(* Logix 5000 project; controller _GigaDiscovery vendor 1 type 14 code 244 rev 35.11; software revision 35.03; part 15 of 23 *)
(* tags used below, declared in another part *)
   Brake_Delay : TIMER;
   Os : DINT;
   Timer_Loc : TIMER[50];
   All_Rack_Closed_Mem : BOOL;
   All_RESTRAINTS_Opened : BOOL;
   DC_Field_Motor_7 : UDT_CROUT;   // DC Field Motor 7 Gondola Contactor -Q16101E -Q16103E
   DC_Field_Pylon_Motors : UDT_CROUT;   // DC Field Pylon Motors Contactor -Q10101E -Q10103E
   Enable_to_Start : UDT_CROUT;   // Abilitazione allo start QC8011E QC8013E
   Girella_Field_Actuate_During_Inactivity : BOOL;
   Gondola_Drive_Enable : UDT_CROUT;   // Gondola Drive Ch1-Ch2 Start Enable Contactors -Q16105E -Q16107E
   I_EStop_Pb_OCC1 : UDT_DCI_STOP_TEST;   // +OCC E-stop -S30301F
   I_EStop_Pb_OCC2 : UDT_DCI_STOP_TEST;   // +OCC2 E-Stop -S28502F
   I_Gondola_Home_Position : BOOL;   // Gondola Home Position -B40002I -B40007I
   I_OCC2_Disable : UDT_DCM;   // OCC 2 CONTROL DISABLE Page 310
   I_OCC_LockOut_Motion : UDT_DCM;   // OCC -Lockout Motion -Q31203E
   I_OCC_Operator_Enable_Key : BOOL;   // OCC Console Enabled -S30305F
   I_Platform_Line_Unlock_Pressure_Switch : BOOL;   // Unlock Platform Line Pressure Switch -S22006B
   I_Platform_Opened : UDT_DCM;   // Platform Opened RFID Series -Q23801J -Q23807J
   I_Platform_Pressure_on_Close_Circuit : BOOL;   // Platform Maximum Closing Pressure -S21510B
   No_Sfty : Std_to_Sfty;
   O_Brake_Pylon_Motor : BOOL;
   Platform_Close_Cycle : Sequencer;
   Platform_Fbk_Valv_Open : BOOL;   // Platform Open Main Valve Limit Switch -B21905I
   Platform_Open_Permissive : Permissive;
   PltaformOpeneded_CycleComplete : BOOL;   // Rilevazione Piattaforme aperte con ciclo Completato
   ProofTest_Req : BOOL;
   Pylon_Field_Actuate_During_Inactivity : BOOL;
   Pylon_Home_Position : UDT_DCM;   // Home position Pylon -B26002I -B26007I
   Pylon_Start_Drive_1_2 : UDT_CROUT;   // Pylon Start Drive 1 - 2 Contactors -Q9002H -Q9004H -Q10202G
   Pylon_Start_Drive_3_4 : UDT_CROUT;   // Pylon Start Drive 3 - 4 Contactors -Q9005H -Q9007H -Q12202G
   Pylon_Start_Drive_5_6 : UDT_CROUT;   // Pylon Start Drive 5 - 6 Contactors -Q9009E -Q9011E4 -Q14202G -Q14202G
   RESTRAINTS_ChA_Open_Memory : BOOL;
   RESTRAINTS_ChB_Open_Memory : BOOL;
   Restraints_Cycle : Sequencer;
   RESTRAINTS_Open_Cycle_Ok : BOOL;
   RESTRAINTS_OpenComand : BOOL;   // Steps 01, 02, 03, 04
   RESTRAINTS_Rack : LapBar_Racks[41];
   RESTRAINTS_Sector : LapBars_Sector[9];
   Start_Autom_Cycle : Sequencer;
   Start_Stop_Cycle : Sequencer;
   Start_TOF : TIMER;
   Valve_Proof_Test_Cycle : Sequencer;
   Valve_Proof_Test_Ok : BOOL;
   Valve_Test_AOI : Sequencer_AOI;
(* S_Cycles, continued *)

ROUTINE _05_Valve_Proof_Test   (* ladder *)
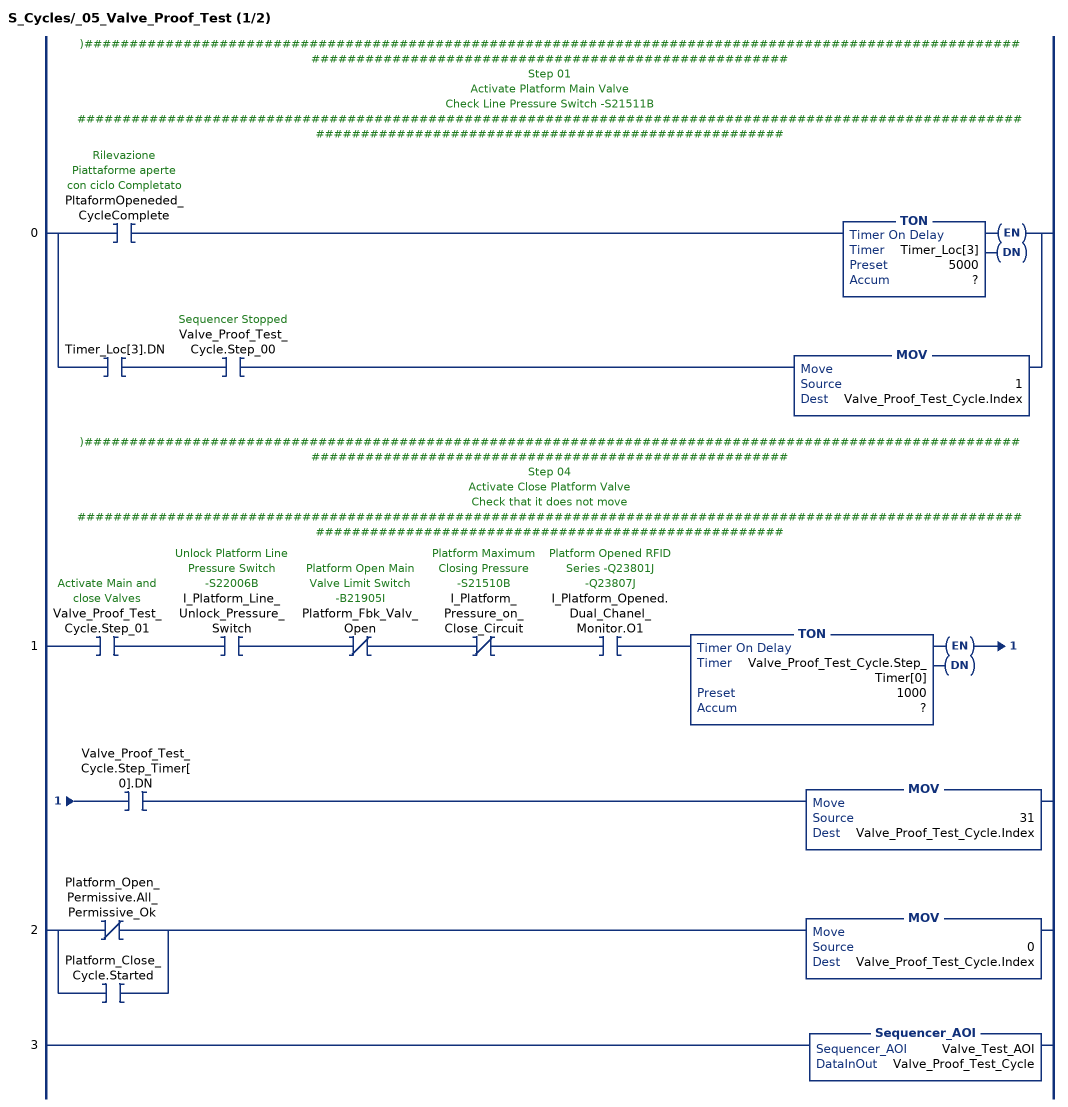
   // )#############################################################################################################################################################
   // Step 01
   // Activate Platform Main Valve
   // Check Line Pressure Switch -S21511B
   // #############################################################################################################################################################
   0: [XIC(PltaformOpeneded_CycleComplete) TON(Timer_Loc[3],?,?) ,XIC(Timer_Loc[3].DN) XIC(Valve_Proof_Test_Cycle.Step_00) MOV(1,Valve_Proof_Test_Cycle.Index) ];
   // )#############################################################################################################################################################
   // Step 04
   // Activate Close Platform Valve
   // Check that it does not move
   // #############################################################################################################################################################
   1: XIC(Valve_Proof_Test_Cycle.Step_01)XIC(I_Platform_Line_Unlock_Pressure_Switch)XIO(Platform_Fbk_Valv_Open)XIO(I_Platform_Pressure_on_Close_Circuit)XIC(I_Platform_Opened.Dual_Chanel_Monitor.O1)TON(Valve_Proof_Test_Cycle.Step_Timer[0],?,?)XIC(Valve_Proof_Test_Cycle.Step_Timer[0].DN)MOV(31,Valve_Proof_Test_Cycle.Index);
   2: [XIO(Platform_Open_Permissive.All_Permissive_Ok) ,XIC(Platform_Close_Cycle.Started) ]MOV(0,Valve_Proof_Test_Cycle.Index);
   3: Sequencer_AOI(Valve_Test_AOI,Valve_Proof_Test_Cycle);
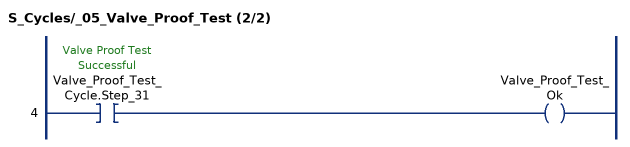
   4: XIC(Valve_Proof_Test_Cycle.Step_31)OTE(Valve_Proof_Test_Ok);
END_ROUTINE

ROUTINE _06_Sensor_Memories   (* ladder *)
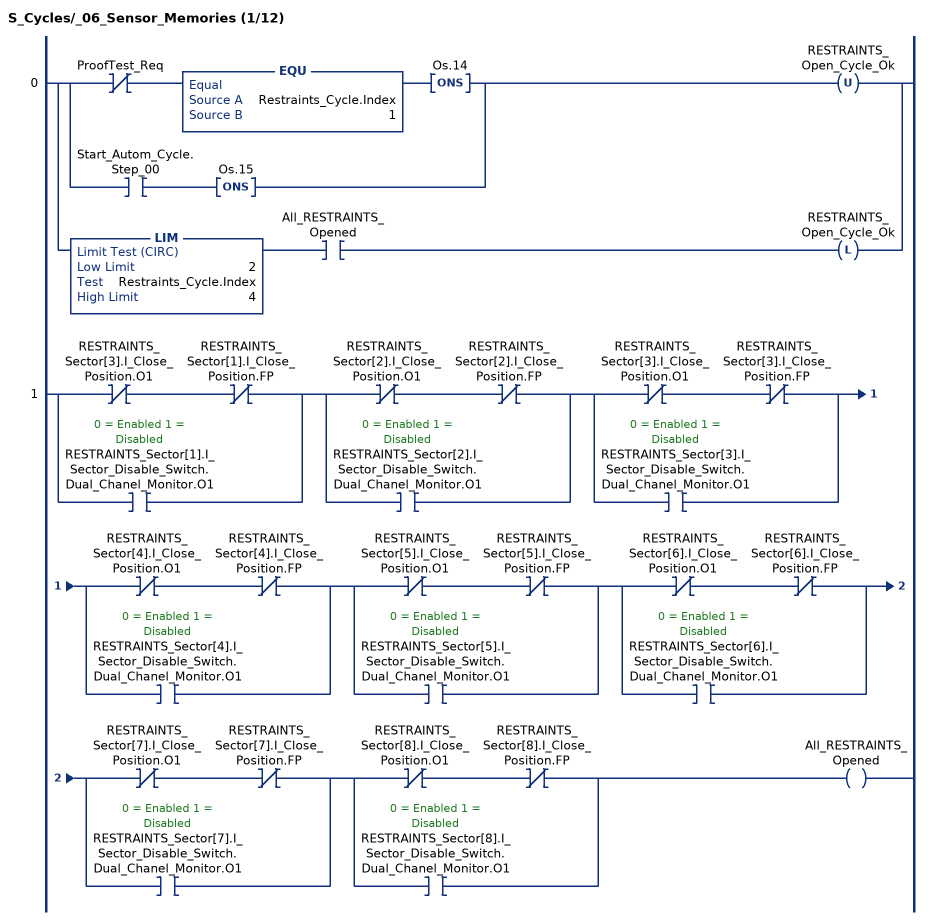
   0: [[XIO(ProofTest_Req) EQU(Restraints_Cycle.Index,1) ONS(Os.14) ,XIC(Start_Autom_Cycle.Step_00) ONS(Os.15) ] OTU(RESTRAINTS_Open_Cycle_Ok) ,LIM(2,Restraints_Cycle.Index,4) XIC(All_RESTRAINTS_Opened) OTL(RESTRAINTS_Open_Cycle_Ok) ];
   1: [XIO(RESTRAINTS_Sector[3].I_Close_Position.O1) XIO(RESTRAINTS_Sector[1].I_Close_Position.FP) ,XIC(RESTRAINTS_Sector[1].I_Sector_Disable_Switch.Dual_Chanel_Monitor.O1) ][XIO(RESTRAINTS_Sector[2].I_Close_Position.O1) XIO(RESTRAINTS_Sector[2].I_Close_Position.FP) ,XIC(RESTRAINTS_Sector[2].I_Sector_Disable_Switch.Dual_Chanel_Monitor.O1) ][XIO(RESTRAINTS_Sector[3].I_Close_Position.O1) XIO(RESTRAINTS_Sector[3].I_Close_Position.FP) ,XIC(RESTRAINTS_Sector[3].I_Sector_Disable_Switch.Dual_Chanel_Monitor.O1) ][XIO(RESTRAINTS_Sector[4].I_Close_Position.O1) XIO(RESTRAINTS_Sector[4].I_Close_Position.FP) ,XIC(RESTRAINTS_Sector[4].I_Sector_Disable_Switch.Dual_Chanel_Monitor.O1) ][XIO(RESTRAINTS_Sector[5].I_Close_Position.O1) XIO(RESTRAINTS_Sector[5].I_Close_Position.FP) ,XIC(RESTRAINTS_Sector[5].I_Sector_Disable_Switch.Dual_Chanel_Monitor.O1) ][XIO(RESTRAINTS_Sector[6].I_Close_Position.O1) XIO(RESTRAINTS_Sector[6].I_Close_Position.FP) ,XIC(RESTRAINTS_Sector[6].I_Sector_Disable_Switch.Dual_Chanel_Monitor.O1) ][XIO(RESTRAINTS_Sector[7].I_Close_Position.O1) XIO(RESTRAINTS_Sector[7].I_Close_Position.FP) ,XIC(RESTRAINTS_Sector[7].I_Sector_Disable_Switch.Dual_Chanel_Monitor.O1) ][XIO(RESTRAINTS_Sector[8].I_Close_Position.O1) XIO(RESTRAINTS_Sector[8].I_Close_Position.FP) ,XIC(RESTRAINTS_Sector[8].I_Sector_Disable_Switch.Dual_Chanel_Monitor.O1) ]OTE(All_RESTRAINTS_Opened);
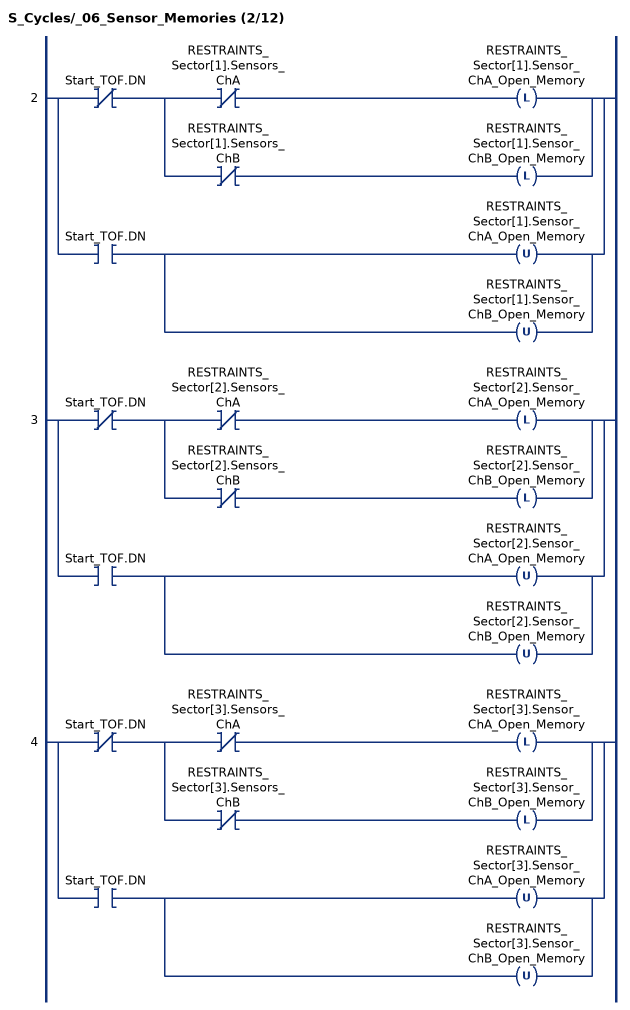
   2: [XIO(Start_TOF.DN) [XIO(RESTRAINTS_Sector[1].Sensors_ChA) OTL(RESTRAINTS_Sector[1].Sensor_ChA_Open_Memory) ,XIO(RESTRAINTS_Sector[1].Sensors_ChB) OTL(RESTRAINTS_Sector[1].Sensor_ChB_Open_Memory) ] ,XIC(Start_TOF.DN) [OTU(RESTRAINTS_Sector[1].Sensor_ChA_Open_Memory) ,OTU(RESTRAINTS_Sector[1].Sensor_ChB_Open_Memory) ] ];
   3: [XIO(Start_TOF.DN) [XIO(RESTRAINTS_Sector[2].Sensors_ChA) OTL(RESTRAINTS_Sector[2].Sensor_ChA_Open_Memory) ,XIO(RESTRAINTS_Sector[2].Sensors_ChB) OTL(RESTRAINTS_Sector[2].Sensor_ChB_Open_Memory) ] ,XIC(Start_TOF.DN) [OTU(RESTRAINTS_Sector[2].Sensor_ChA_Open_Memory) ,OTU(RESTRAINTS_Sector[2].Sensor_ChB_Open_Memory) ] ];
   4: [XIO(Start_TOF.DN) [XIO(RESTRAINTS_Sector[3].Sensors_ChA) OTL(RESTRAINTS_Sector[3].Sensor_ChA_Open_Memory) ,XIO(RESTRAINTS_Sector[3].Sensors_ChB) OTL(RESTRAINTS_Sector[3].Sensor_ChB_Open_Memory) ] ,XIC(Start_TOF.DN) [OTU(RESTRAINTS_Sector[3].Sensor_ChA_Open_Memory) ,OTU(RESTRAINTS_Sector[3].Sensor_ChB_Open_Memory) ] ];
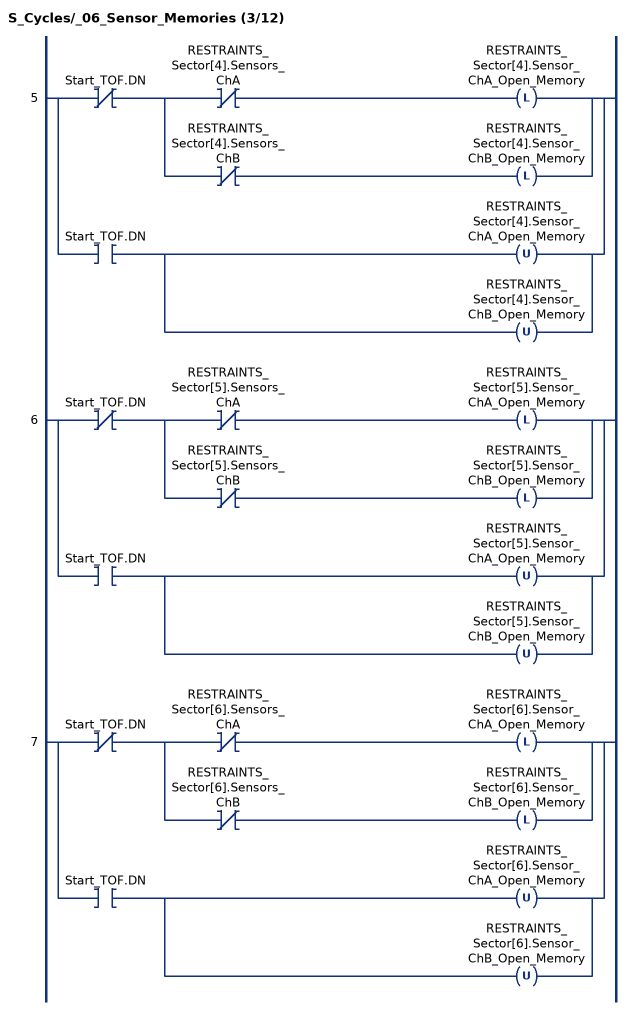
   5: [XIO(Start_TOF.DN) [XIO(RESTRAINTS_Sector[4].Sensors_ChA) OTL(RESTRAINTS_Sector[4].Sensor_ChA_Open_Memory) ,XIO(RESTRAINTS_Sector[4].Sensors_ChB) OTL(RESTRAINTS_Sector[4].Sensor_ChB_Open_Memory) ] ,XIC(Start_TOF.DN) [OTU(RESTRAINTS_Sector[4].Sensor_ChA_Open_Memory) ,OTU(RESTRAINTS_Sector[4].Sensor_ChB_Open_Memory) ] ];
   6: [XIO(Start_TOF.DN) [XIO(RESTRAINTS_Sector[5].Sensors_ChA) OTL(RESTRAINTS_Sector[5].Sensor_ChA_Open_Memory) ,XIO(RESTRAINTS_Sector[5].Sensors_ChB) OTL(RESTRAINTS_Sector[5].Sensor_ChB_Open_Memory) ] ,XIC(Start_TOF.DN) [OTU(RESTRAINTS_Sector[5].Sensor_ChA_Open_Memory) ,OTU(RESTRAINTS_Sector[5].Sensor_ChB_Open_Memory) ] ];
   7: [XIO(Start_TOF.DN) [XIO(RESTRAINTS_Sector[6].Sensors_ChA) OTL(RESTRAINTS_Sector[6].Sensor_ChA_Open_Memory) ,XIO(RESTRAINTS_Sector[6].Sensors_ChB) OTL(RESTRAINTS_Sector[6].Sensor_ChB_Open_Memory) ] ,XIC(Start_TOF.DN) [OTU(RESTRAINTS_Sector[6].Sensor_ChA_Open_Memory) ,OTU(RESTRAINTS_Sector[6].Sensor_ChB_Open_Memory) ] ];
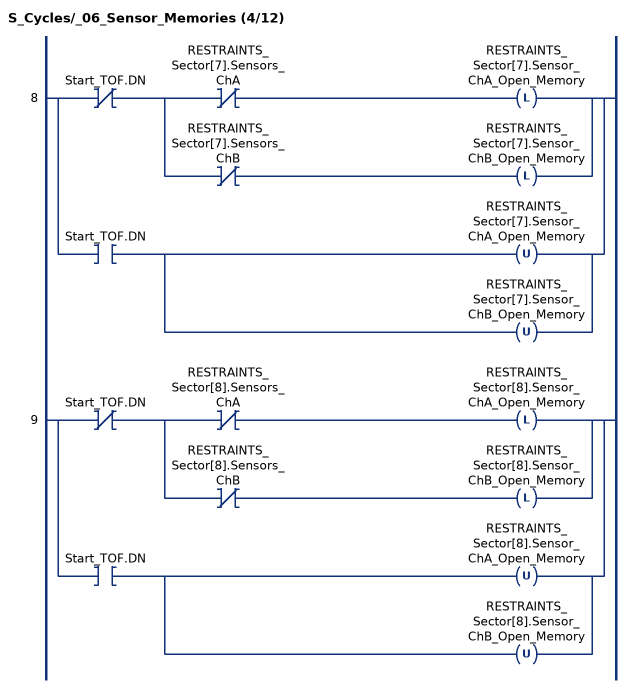
   8: [XIO(Start_TOF.DN) [XIO(RESTRAINTS_Sector[7].Sensors_ChA) OTL(RESTRAINTS_Sector[7].Sensor_ChA_Open_Memory) ,XIO(RESTRAINTS_Sector[7].Sensors_ChB) OTL(RESTRAINTS_Sector[7].Sensor_ChB_Open_Memory) ] ,XIC(Start_TOF.DN) [OTU(RESTRAINTS_Sector[7].Sensor_ChA_Open_Memory) ,OTU(RESTRAINTS_Sector[7].Sensor_ChB_Open_Memory) ] ];
   9: [XIO(Start_TOF.DN) [XIO(RESTRAINTS_Sector[8].Sensors_ChA) OTL(RESTRAINTS_Sector[8].Sensor_ChA_Open_Memory) ,XIO(RESTRAINTS_Sector[8].Sensors_ChB) OTL(RESTRAINTS_Sector[8].Sensor_ChB_Open_Memory) ] ,XIC(Start_TOF.DN) [OTU(RESTRAINTS_Sector[8].Sensor_ChA_Open_Memory) ,OTU(RESTRAINTS_Sector[8].Sensor_ChB_Open_Memory) ] ];
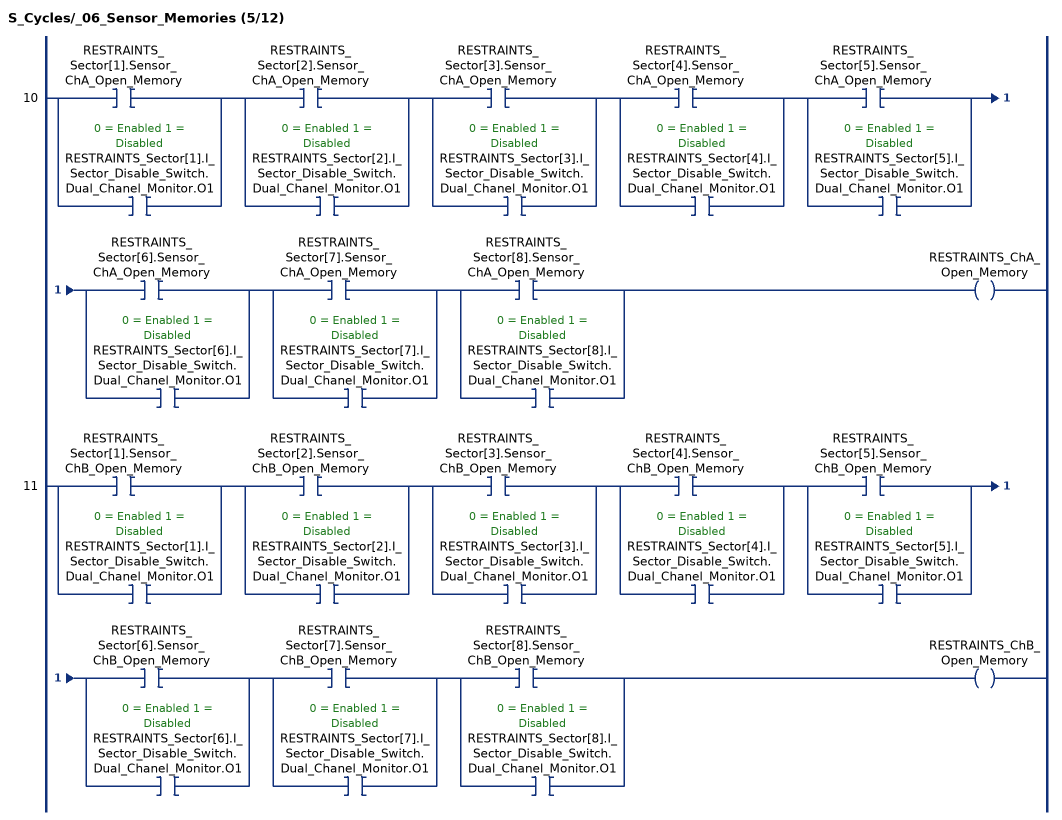
   10: [XIC(RESTRAINTS_Sector[1].Sensor_ChA_Open_Memory) ,XIC(RESTRAINTS_Sector[1].I_Sector_Disable_Switch.Dual_Chanel_Monitor.O1) ][XIC(RESTRAINTS_Sector[2].Sensor_ChA_Open_Memory) ,XIC(RESTRAINTS_Sector[2].I_Sector_Disable_Switch.Dual_Chanel_Monitor.O1) ][XIC(RESTRAINTS_Sector[3].Sensor_ChA_Open_Memory) ,XIC(RESTRAINTS_Sector[3].I_Sector_Disable_Switch.Dual_Chanel_Monitor.O1) ][XIC(RESTRAINTS_Sector[4].Sensor_ChA_Open_Memory) ,XIC(RESTRAINTS_Sector[4].I_Sector_Disable_Switch.Dual_Chanel_Monitor.O1) ][XIC(RESTRAINTS_Sector[5].Sensor_ChA_Open_Memory) ,XIC(RESTRAINTS_Sector[5].I_Sector_Disable_Switch.Dual_Chanel_Monitor.O1) ][XIC(RESTRAINTS_Sector[6].Sensor_ChA_Open_Memory) ,XIC(RESTRAINTS_Sector[6].I_Sector_Disable_Switch.Dual_Chanel_Monitor.O1) ][XIC(RESTRAINTS_Sector[7].Sensor_ChA_Open_Memory) ,XIC(RESTRAINTS_Sector[7].I_Sector_Disable_Switch.Dual_Chanel_Monitor.O1) ][XIC(RESTRAINTS_Sector[8].Sensor_ChA_Open_Memory) ,XIC(RESTRAINTS_Sector[8].I_Sector_Disable_Switch.Dual_Chanel_Monitor.O1) ]OTE(RESTRAINTS_ChA_Open_Memory);
   11: [XIC(RESTRAINTS_Sector[1].Sensor_ChB_Open_Memory) ,XIC(RESTRAINTS_Sector[1].I_Sector_Disable_Switch.Dual_Chanel_Monitor.O1) ][XIC(RESTRAINTS_Sector[2].Sensor_ChB_Open_Memory) ,XIC(RESTRAINTS_Sector[2].I_Sector_Disable_Switch.Dual_Chanel_Monitor.O1) ][XIC(RESTRAINTS_Sector[3].Sensor_ChB_Open_Memory) ,XIC(RESTRAINTS_Sector[3].I_Sector_Disable_Switch.Dual_Chanel_Monitor.O1) ][XIC(RESTRAINTS_Sector[4].Sensor_ChB_Open_Memory) ,XIC(RESTRAINTS_Sector[4].I_Sector_Disable_Switch.Dual_Chanel_Monitor.O1) ][XIC(RESTRAINTS_Sector[5].Sensor_ChB_Open_Memory) ,XIC(RESTRAINTS_Sector[5].I_Sector_Disable_Switch.Dual_Chanel_Monitor.O1) ][XIC(RESTRAINTS_Sector[6].Sensor_ChB_Open_Memory) ,XIC(RESTRAINTS_Sector[6].I_Sector_Disable_Switch.Dual_Chanel_Monitor.O1) ][XIC(RESTRAINTS_Sector[7].Sensor_ChB_Open_Memory) ,XIC(RESTRAINTS_Sector[7].I_Sector_Disable_Switch.Dual_Chanel_Monitor.O1) ][XIC(RESTRAINTS_Sector[8].Sensor_ChB_Open_Memory) ,XIC(RESTRAINTS_Sector[8].I_Sector_Disable_Switch.Dual_Chanel_Monitor.O1) ]OTE(RESTRAINTS_ChB_Open_Memory);
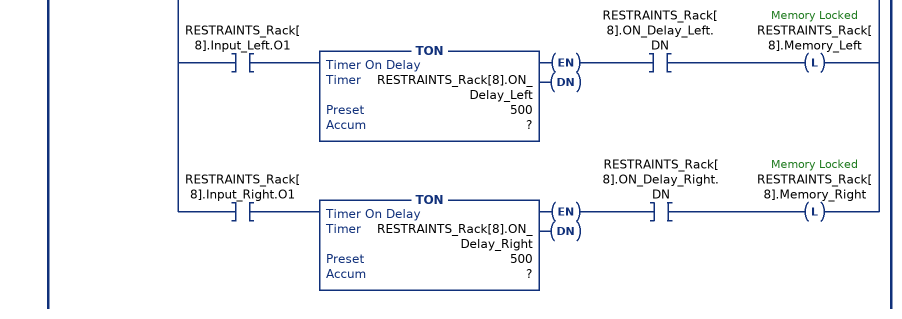
   12: XIC(Restraints_Cycle.Step_22)[XIC(RESTRAINTS_Rack[1].Input_Left.O1) TON(RESTRAINTS_Rack[1].ON_Delay_Left,?,?) XIC(RESTRAINTS_Rack[1].ON_Delay_Left.DN) OTL(RESTRAINTS_Rack[1].Memory_Left) ,XIC(RESTRAINTS_Rack[1].Input_Right.O1) TON(RESTRAINTS_Rack[1].ON_Delay_Right,?,?) XIC(RESTRAINTS_Rack[1].ON_Delay_Right.DN) OTL(RESTRAINTS_Rack[1].Memory_Right) ,XIC(RESTRAINTS_Rack[2].Input_Left.O1) TON(RESTRAINTS_Rack[2].ON_Delay_Left,?,?) XIC(RESTRAINTS_Rack[2].ON_Delay_Left.DN) OTL(RESTRAINTS_Rack[2].Memory_Left) ,XIC(RESTRAINTS_Rack[2].Input_Right.O1) TON(RESTRAINTS_Rack[2].ON_Delay_Right,?,?) XIC(RESTRAINTS_Rack[2].ON_Delay_Right.DN) OTL(RESTRAINTS_Rack[2].Memory_Right) ,XIC(RESTRAINTS_Rack[3].Input_Left.O1) TON(RESTRAINTS_Rack[3].ON_Delay_Left,?,?) XIC(RESTRAINTS_Rack[3].ON_Delay_Left.DN) OTL(RESTRAINTS_Rack[3].Memory_Left) ,XIC(RESTRAINTS_Rack[3].Input_Right.O1) TON(RESTRAINTS_Rack[3].ON_Delay_Right,?,?) XIC(RESTRAINTS_Rack[3].ON_Delay_Right.DN) OTL(RESTRAINTS_Rack[3].Memory_Right) ,XIC(RESTRAINTS_Rack[4].Input_Left.O1) TON(RESTRAINTS_Rack[4].ON_Delay_Left,?,?) XIC(RESTRAINTS_Rack[4].ON_Delay_Left.DN) OTL(RESTRAINTS_Rack[4].Memory_Left) ,XIC(RESTRAINTS_Rack[4].Input_Right.O1) TON(RESTRAINTS_Rack[4].ON_Delay_Right,?,?) XIC(RESTRAINTS_Rack[4].ON_Delay_Right.DN) OTL(RESTRAINTS_Rack[4].Memory_Right) ,XIC(RESTRAINTS_Rack[5].Input_Left.O1) TON(RESTRAINTS_Rack[5].ON_Delay_Left,?,?) XIC(RESTRAINTS_Rack[5].ON_Delay_Left.DN) OTL(RESTRAINTS_Rack[5].Memory_Left) ,XIC(RESTRAINTS_Rack[5].Input_Right.O1) TON(RESTRAINTS_Rack[5].ON_Delay_Right,?,?) XIC(RESTRAINTS_Rack[5].ON_Delay_Right.DN) OTL(RESTRAINTS_Rack[5].Memory_Right) ,XIC(RESTRAINTS_Rack[6].Input_Left.O1) TON(RESTRAINTS_Rack[6].ON_Delay_Left,?,?) XIC(RESTRAINTS_Rack[6].ON_Delay_Left.DN) OTL(RESTRAINTS_Rack[6].Memory_Left) ,XIC(RESTRAINTS_Rack[6].Input_Right.O1) TON(RESTRAINTS_Rack[6].ON_Delay_Right,?,?) XIC(RESTRAINTS_Rack[6].ON_Delay_Right.DN) OTL(RESTRAINTS_Rack[6].Memory_Right) ,XIC(RESTRAINTS_Rack[7].Input_Left.O1) TON(RESTRAINTS_Rack[7].ON_Delay_Left,?,?) XIC(RESTRAINTS_Rack[7].ON_Delay_Left.DN) OTL(RESTRAINTS_Rack[7].Memory_Left) ,XIC(RESTRAINTS_Rack[7].Input_Right.O1) TON(RESTRAINTS_Rack[7].ON_Delay_Right,?,?) XIC(RESTRAINTS_Rack[7].ON_Delay_Right.DN) OTL(RESTRAINTS_Rack[7].Memory_Right) ,XIC(RESTRAINTS_Rack[8].Input_Left.O1) TON(RESTRAINTS_Rack[8].ON_Delay_Left,?,?) XIC(RESTRAINTS_Rack[8].ON_Delay_Left.DN) OTL(RESTRAINTS_Rack[8].Memory_Left) ,XIC(RESTRAINTS_Rack[8].Input_Right.O1) TON(RESTRAINTS_Rack[8].ON_Delay_Right,?,?) XIC(RESTRAINTS_Rack[8].ON_Delay_Right.DN) OTL(RESTRAINTS_Rack[8].Memory_Right) ];
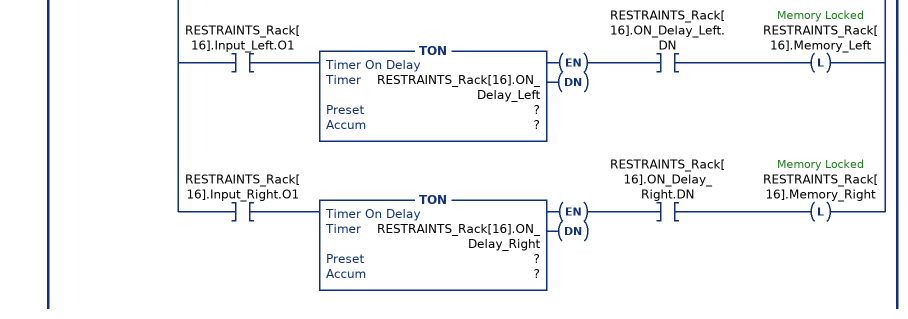
   13: XIC(Restraints_Cycle.Step_22)[XIC(RESTRAINTS_Rack[9].Input_Left.O1) TON(RESTRAINTS_Rack[9].ON_Delay_Left,?,?) XIC(RESTRAINTS_Rack[9].ON_Delay_Left.DN) OTL(RESTRAINTS_Rack[9].Memory_Left) ,XIC(RESTRAINTS_Rack[9].Input_Right.O1) TON(RESTRAINTS_Rack[9].ON_Delay_Right,?,?) XIC(RESTRAINTS_Rack[9].ON_Delay_Right.DN) OTL(RESTRAINTS_Rack[9].Memory_Right) ,XIC(RESTRAINTS_Rack[10].Input_Left.O1) TON(RESTRAINTS_Rack[10].ON_Delay_Left,?,?) XIC(RESTRAINTS_Rack[10].ON_Delay_Left.DN) OTL(RESTRAINTS_Rack[10].Memory_Left) ,XIC(RESTRAINTS_Rack[10].Input_Right.O1) TON(RESTRAINTS_Rack[10].ON_Delay_Right,?,?) XIC(RESTRAINTS_Rack[10].ON_Delay_Right.DN) OTL(RESTRAINTS_Rack[10].Memory_Right) ,XIC(RESTRAINTS_Rack[11].Input_Left.O1) TON(RESTRAINTS_Rack[11].ON_Delay_Left,?,?) XIC(RESTRAINTS_Rack[11].ON_Delay_Left.DN) OTL(RESTRAINTS_Rack[11].Memory_Left) ,XIC(RESTRAINTS_Rack[11].Input_Right.O1) TON(RESTRAINTS_Rack[11].ON_Delay_Right,?,?) XIC(RESTRAINTS_Rack[11].ON_Delay_Right.DN) OTL(RESTRAINTS_Rack[11].Memory_Right) ,XIC(RESTRAINTS_Rack[12].Input_Left.O1) TON(RESTRAINTS_Rack[12].ON_Delay_Left,?,?) XIC(RESTRAINTS_Rack[12].ON_Delay_Left.DN) OTL(RESTRAINTS_Rack[12].Memory_Left) ,XIC(RESTRAINTS_Rack[12].Input_Right.O1) TON(RESTRAINTS_Rack[12].ON_Delay_Right,?,?) XIC(RESTRAINTS_Rack[12].ON_Delay_Right.DN) OTL(RESTRAINTS_Rack[12].Memory_Right) ,XIC(RESTRAINTS_Rack[13].Input_Left.O1) TON(RESTRAINTS_Rack[13].ON_Delay_Left,?,?) XIC(RESTRAINTS_Rack[13].ON_Delay_Left.DN) OTL(RESTRAINTS_Rack[13].Memory_Left) ,XIC(RESTRAINTS_Rack[13].Input_Right.O1) TON(RESTRAINTS_Rack[13].ON_Delay_Right,?,?) XIC(RESTRAINTS_Rack[13].ON_Delay_Right.DN) OTL(RESTRAINTS_Rack[13].Memory_Right) ,XIC(RESTRAINTS_Rack[14].Input_Left.O1) TON(RESTRAINTS_Rack[14].ON_Delay_Left,?,?) XIC(RESTRAINTS_Rack[14].ON_Delay_Left.DN) OTL(RESTRAINTS_Rack[14].Memory_Left) ,XIC(RESTRAINTS_Rack[14].Input_Right.O1) TON(RESTRAINTS_Rack[14].ON_Delay_Right,?,?) XIC(RESTRAINTS_Rack[14].ON_Delay_Right.DN) OTL(RESTRAINTS_Rack[14].Memory_Right) ,XIC(RESTRAINTS_Rack[15].Input_Left.O1) TON(RESTRAINTS_Rack[15].ON_Delay_Left,?,?) XIC(RESTRAINTS_Rack[15].ON_Delay_Left.DN) OTL(RESTRAINTS_Rack[15].Memory_Left) ,XIC(RESTRAINTS_Rack[15].Input_Right.O1) TON(RESTRAINTS_Rack[15].ON_Delay_Right,?,?) XIC(RESTRAINTS_Rack[15].ON_Delay_Right.DN) OTL(RESTRAINTS_Rack[15].Memory_Right) ,XIC(RESTRAINTS_Rack[16].Input_Left.O1) TON(RESTRAINTS_Rack[16].ON_Delay_Left,?,?) XIC(RESTRAINTS_Rack[16].ON_Delay_Left.DN) OTL(RESTRAINTS_Rack[16].Memory_Left) ,XIC(RESTRAINTS_Rack[16].Input_Right.O1) TON(RESTRAINTS_Rack[16].ON_Delay_Right,?,?) XIC(RESTRAINTS_Rack[16].ON_Delay_Right.DN) OTL(RESTRAINTS_Rack[16].Memory_Right) ];